REGION Network 4: Run IGG Sea Water P301-CV311-CV322
   // Changed to 560 from 580
   RUNG wire#powerrail
      { S7_Templates := "SrcType := Int" } GE_Contact(in1 := "100_GCU_AUTO_SEQ_DB".CRNT_STEP, in2 := 50)
      { S7_Templates := "SrcType := Int" } LE_Contact(in1 := "100_GCU_AUTO_SEQ_DB".CRNT_STEP, in2 := 560)
      wire#w1
      Contact( "51_SLAVE_STATUS".CV322_OPN )
      Contact( "51_SLAVE_STATUS"."CV-321_CLSD" )
      Coil( "56_SLAVE_CMNDS".OPEN_CV311 )
   END_RUNG
   RUNG wire#powerrail
      I_Contact( "10_DI_DATA".E_400_STPD )
      I_Contact( "10_DI_DATA".E_400_SHTDN )
   END_RUNG wire#w1
   RUNG wire#w1
      Coil( "56_SLAVE_CMNDS".OPEN_CV322 )
   END_RUNG
   RUNG wire#w1
      Contact( "51_SLAVE_STATUS".CV311_OPN )
      Contact( "51_SLAVE_STATUS".CV322_OPN )
      Coil( "56_SLAVE_CMNDS".RUN_P301 )
   END_RUNG
   // the same network as SCL:
   #_w1 := (("100_GCU_AUTO_SEQ_DB".CRNT_STEP >= 50) AND ("100_GCU_AUTO_SEQ_DB".CRNT_STEP <= 560)) OR (NOT "10_DI_DATA".E_400_STPD AND NOT "10_DI_DATA".E_400_SHTDN);
   "56_SLAVE_CMNDS".OPEN_CV311 := #_w1 AND "51_SLAVE_STATUS".CV322_OPN AND "51_SLAVE_STATUS"."CV-321_CLSD";
   "56_SLAVE_CMNDS".OPEN_CV322 := #_w1;
   "56_SLAVE_CMNDS".RUN_P301 := #_w1 AND "51_SLAVE_STATUS".CV311_OPN AND "51_SLAVE_STATUS".CV322_OPN;
END_REGION

REGION Network 5: Q136.0 - Fresh Water Fill Valve Control(CV358)
   // True = RUN, False = NOT
   RUNG wire#powerrail
      { S7_Templates := "SrcType := Int" } GE_Contact(in1 := "100_GCU_AUTO_SEQ_DB".CRNT_STEP, in2 := 90)
      { S7_Templates := "SrcType := Int" } LT_Contact(in1 := "100_GCU_AUTO_SEQ_DB".CRNT_STEP, in2 := 200)
      wire#w1
      Coil( "14_DQ_DATA".CV_358 )
   END_RUNG
   RUNG wire#powerrail
      Contact( "108_GCU_TNK_REFILL_SEQ_DB".OPEN_CV358 )
   END_RUNG wire#w1
   RUNG wire#powerrail
      Contact( "110_GCU_TNK_FLUSH_SEQ_DB".OPEN_CV358 )
   END_RUNG wire#w1
   // the same network as SCL:
   "14_DQ_DATA".CV_358 := (("100_GCU_AUTO_SEQ_DB".CRNT_STEP >= 90) AND ("100_GCU_AUTO_SEQ_DB".CRNT_STEP < 200)) OR "108_GCU_TNK_REFILL_SEQ_DB".OPEN_CV358 OR "110_GCU_TNK_FLUSH_SEQ_DB".OPEN_CV358;
END_REGION

REGION Network 6: Q136.1 - Waste Water Drain Valve Control (CV341)
   // True = Close, False = Open    Condition added to avoid back filling the GCU through common drain on Bordeira
   RUNG wire#powerrail
      { S7_Templates := "SrcType := Int" } GE_Contact(in1 := "100_GCU_AUTO_SEQ_DB".CRNT_STEP, in2 := 60)
      { S7_Templates := "SrcType := Int" } LT_Contact(in1 := "100_GCU_AUTO_SEQ_DB".CRNT_STEP, in2 := 570)
      wire#w1
      Coil( "14_DQ_DATA".CV_341 )
   END_RUNG
   RUNG wire#powerrail
      I_Contact( "51_SLAVE_STATUS".CV311_CLSD )
      Contact( "AlwaysTRUE" )
   END_RUNG wire#w1
   // the same network as SCL:
   "14_DQ_DATA".CV_341 := (("100_GCU_AUTO_SEQ_DB".CRNT_STEP >= 60) AND ("100_GCU_AUTO_SEQ_DB".CRNT_STEP < 570)) OR (NOT "51_SLAVE_STATUS".CV311_CLSD AND "AlwaysTRUE");
END_REGION

REGION Network 7: Q136.2 - Block Valve 1 Control (CV407) +++Control By BWTS+++
   // True = RUN, False = NOT
END_REGION

REGION Network 8: Q136.3 - Bleed Valve Control (CV409) +++Control By BWTS+++
   // True = OPEN, False = CLOSE
END_REGION

REGION Network 9: Q136.4 - Block Valve 2 Control (CV411) +++Control By BWTS+++
   // True = OPEN, False = CLOSE
END_REGION

REGION Network 10: Q136.5 - Ambient Air Valve Control (CV441)
   // True = CLOSE, False = OPEN        STOP bits are redundant.
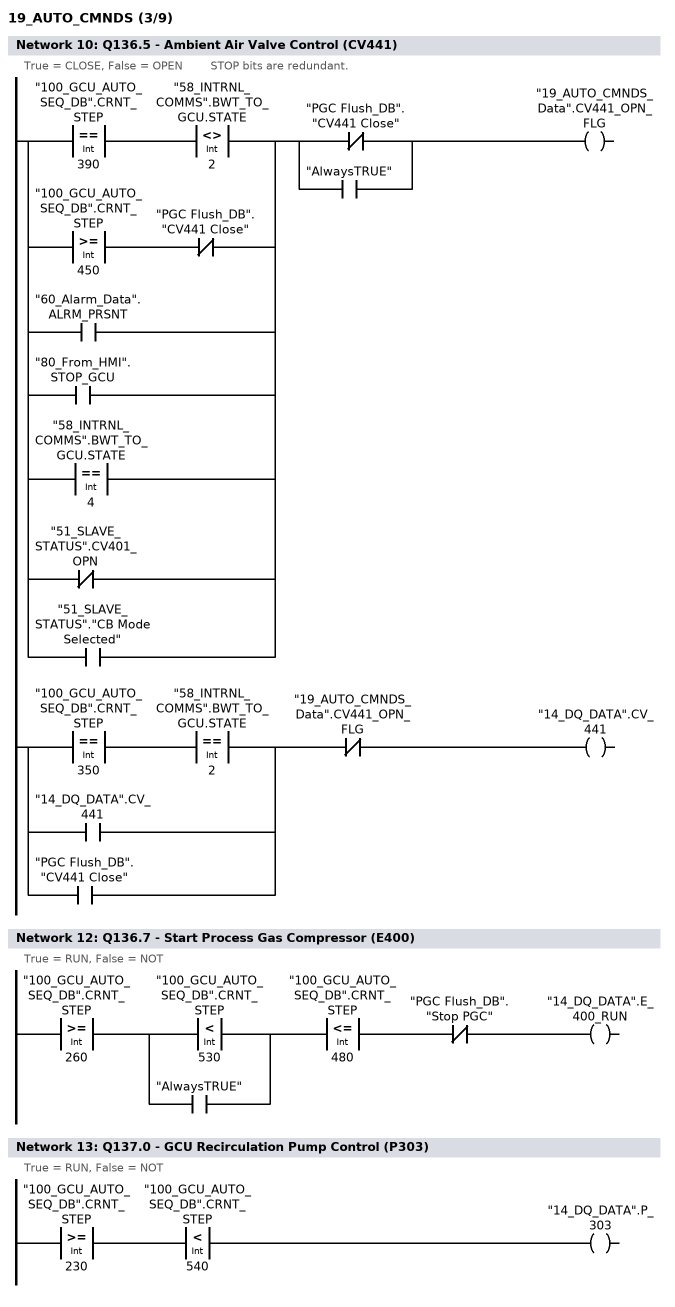
   RUNG wire#powerrail
      { S7_Templates := "SrcType := Int" } EQ_Contact(in1 := "100_GCU_AUTO_SEQ_DB".CRNT_STEP, in2 := 390)
      { S7_Templates := "SrcType := Int" } NE_Contact(in1 := "58_INTRNL_COMMS".BWT_TO_GCU.STATE, in2 := 2)
      wire#w1
      I_Contact( "PGC Flush_DB"."CV441 Close" )
      wire#w2
      Coil( "19_AUTO_CMNDS_Data".CV441_OPN_FLG )
   END_RUNG
   RUNG wire#powerrail
      { S7_Templates := "SrcType := Int" } GE_Contact(in1 := "100_GCU_AUTO_SEQ_DB".CRNT_STEP, in2 := 450)
      I_Contact( "PGC Flush_DB"."CV441 Close" )
   END_RUNG wire#w1
   RUNG wire#powerrail
      Contact( "60_Alarm_Data".ALRM_PRSNT )
   END_RUNG wire#w1
   RUNG wire#powerrail
      Contact( "80_From_HMI".STOP_GCU )
   END_RUNG wire#w1
   RUNG wire#powerrail
      { S7_Templates := "SrcType := Int" } EQ_Contact(in1 := "58_INTRNL_COMMS".BWT_TO_GCU.STATE, in2 := 4)
   END_RUNG wire#w1
   RUNG wire#powerrail
      I_Contact( "51_SLAVE_STATUS".CV401_OPN )
   END_RUNG wire#w1
   RUNG wire#powerrail
      Contact( "51_SLAVE_STATUS"."CB Mode Selected" )
   END_RUNG wire#w1
   RUNG wire#w1
      Contact( "AlwaysTRUE" )
   END_RUNG wire#w2
   RUNG wire#powerrail
      { S7_Templates := "SrcType := Int" } EQ_Contact(in1 := "100_GCU_AUTO_SEQ_DB".CRNT_STEP, in2 := 350)
      { S7_Templates := "SrcType := Int" } EQ_Contact(in1 := "58_INTRNL_COMMS".BWT_TO_GCU.STATE, in2 := 2)
      wire#w3
      I_Contact( "19_AUTO_CMNDS_Data".CV441_OPN_FLG )
      Coil( "14_DQ_DATA".CV_441 )
   END_RUNG
   RUNG wire#powerrail
      Contact( "14_DQ_DATA".CV_441 )
   END_RUNG wire#w3
   RUNG wire#powerrail
      Contact( "PGC Flush_DB"."CV441 Close" )
   END_RUNG wire#w3
   // the same network as SCL:
   "19_AUTO_CMNDS_Data".CV441_OPN_FLG := ((("100_GCU_AUTO_SEQ_DB".CRNT_STEP = 390) AND ("58_INTRNL_COMMS".BWT_TO_GCU.STATE <> 2)) OR (("100_GCU_AUTO_SEQ_DB".CRNT_STEP >= 450) AND NOT "PGC Flush_DB"."CV441 Close") OR "60_Alarm_Data".ALRM_PRSNT OR "80_From_HMI".STOP_GCU OR ("58_INTRNL_COMMS".BWT_TO_GCU.STATE = 4) OR NOT "51_SLAVE_STATUS".CV401_OPN OR "51_SLAVE_STATUS"."CB Mode Selected") AND (NOT "PGC Flush_DB"."CV441 Close" OR "AlwaysTRUE");
   "14_DQ_DATA".CV_441 := ((("100_GCU_AUTO_SEQ_DB".CRNT_STEP = 350) AND ("58_INTRNL_COMMS".BWT_TO_GCU.STATE = 2)) OR "14_DQ_DATA".CV_441 OR "PGC Flush_DB"."CV441 Close") AND NOT "19_AUTO_CMNDS_Data".CV441_OPN_FLG;
END_REGION

REGION Network 11: Q136.6 - Main Gas to Deck Valve Control (CV406) +++Control By BWTS+++
   // True = RUN, False = NOT
END_REGION

REGION Network 12: Q136.7 - Start Process Gas Compressor (E400)
   // True = RUN, False = NOT
   RUNG wire#powerrail
      { S7_Templates := "SrcType := Int" } GE_Contact(in1 := "100_GCU_AUTO_SEQ_DB".CRNT_STEP, in2 := 260)
      wire#w1
      { S7_Templates := "SrcType := Int" } LT_Contact(in1 := "100_GCU_AUTO_SEQ_DB".CRNT_STEP, in2 := 530)
      wire#w2
      { S7_Templates := "SrcType := Int" } LE_Contact(in1 := "100_GCU_AUTO_SEQ_DB".CRNT_STEP, in2 := 480)
      I_Contact( "PGC Flush_DB"."Stop PGC" )
      Coil( "14_DQ_DATA".E_400_RUN )
   END_RUNG
   RUNG wire#w1
      Contact( "AlwaysTRUE" )
   END_RUNG wire#w2
   // the same network as SCL:
   "14_DQ_DATA".E_400_RUN := ("100_GCU_AUTO_SEQ_DB".CRNT_STEP >= 260) AND (("100_GCU_AUTO_SEQ_DB".CRNT_STEP < 530) OR "AlwaysTRUE") AND ("100_GCU_AUTO_SEQ_DB".CRNT_STEP <= 480) AND NOT "PGC Flush_DB"."Stop PGC";
END_REGION

REGION Network 13: Q137.0 - GCU Recirculation Pump Control (P303)
   // True = RUN, False = NOT
   RUNG wire#powerrail
      { S7_Templates := "SrcType := Int" } GE_Contact(in1 := "100_GCU_AUTO_SEQ_DB".CRNT_STEP, in2 := 230)
      { S7_Templates := "SrcType := Int" } LT_Contact(in1 := "100_GCU_AUTO_SEQ_DB".CRNT_STEP, in2 := 540)
      Coil( "14_DQ_DATA".P_303 )
   END_RUNG
   // the same network as SCL:
   "14_DQ_DATA".P_303 := ("100_GCU_AUTO_SEQ_DB".CRNT_STEP >= 230) AND ("100_GCU_AUTO_SEQ_DB".CRNT_STEP < 540);
END_REGION

REGION Network 14: Q137.1 - GCU Booster Pump Control (P304)
   // True = ALARM, False = NOT
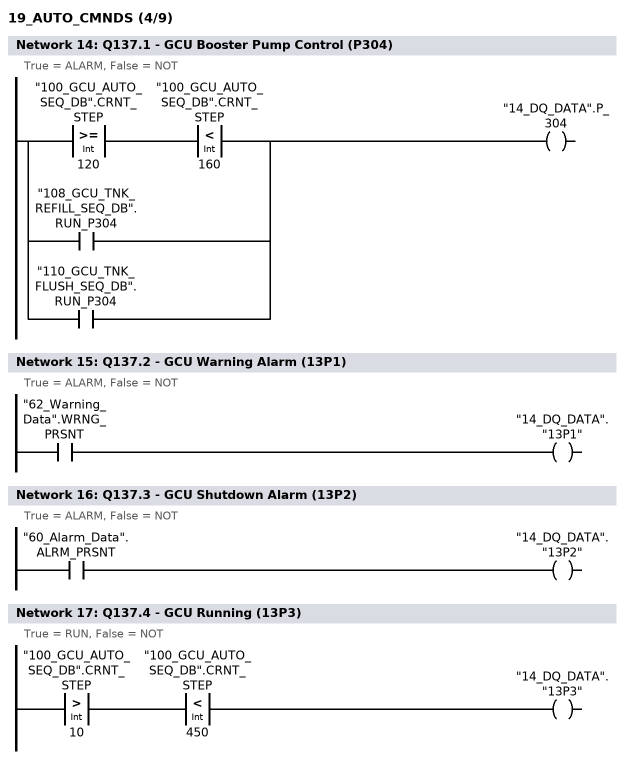
   RUNG wire#powerrail
      { S7_Templates := "SrcType := Int" } GE_Contact(in1 := "100_GCU_AUTO_SEQ_DB".CRNT_STEP, in2 := 120)
      { S7_Templates := "SrcType := Int" } LT_Contact(in1 := "100_GCU_AUTO_SEQ_DB".CRNT_STEP, in2 := 160)
      wire#w1
      Coil( "14_DQ_DATA".P_304 )
   END_RUNG
   RUNG wire#powerrail
      Contact( "108_GCU_TNK_REFILL_SEQ_DB".RUN_P304 )
   END_RUNG wire#w1
   RUNG wire#powerrail
      Contact( "110_GCU_TNK_FLUSH_SEQ_DB".RUN_P304 )
   END_RUNG wire#w1
   // the same network as SCL:
   "14_DQ_DATA".P_304 := (("100_GCU_AUTO_SEQ_DB".CRNT_STEP >= 120) AND ("100_GCU_AUTO_SEQ_DB".CRNT_STEP < 160)) OR "108_GCU_TNK_REFILL_SEQ_DB".RUN_P304 OR "110_GCU_TNK_FLUSH_SEQ_DB".RUN_P304;
END_REGION

REGION Network 15: Q137.2 - GCU Warning Alarm (13P1)
   // True = ALARM, False = NOT
   RUNG wire#powerrail
      Contact( "62_Warning_Data".WRNG_PRSNT )
      Coil( "14_DQ_DATA"."13P1" )
   END_RUNG
   // the same network as SCL:
   "14_DQ_DATA"."13P1" := "62_Warning_Data".WRNG_PRSNT;
END_REGION

REGION Network 16: Q137.3 - GCU Shutdown Alarm (13P2)
   // True = ALARM, False = NOT
   RUNG wire#powerrail
      Contact( "60_Alarm_Data".ALRM_PRSNT )
      Coil( "14_DQ_DATA"."13P2" )
   END_RUNG
   // the same network as SCL:
   "14_DQ_DATA"."13P2" := "60_Alarm_Data".ALRM_PRSNT;
END_REGION

REGION Network 17: Q137.4 - GCU Running (13P3)
   // True = RUN, False = NOT
   RUNG wire#powerrail
      { S7_Templates := "SrcType := Int" } GT_Contact(in1 := "100_GCU_AUTO_SEQ_DB".CRNT_STEP, in2 := 10)
      { S7_Templates := "SrcType := Int" } LT_Contact(in1 := "100_GCU_AUTO_SEQ_DB".CRNT_STEP, in2 := 450)
      Coil( "14_DQ_DATA"."13P3" )
   END_RUNG
   // the same network as SCL:
   "14_DQ_DATA"."13P3" := ("100_GCU_AUTO_SEQ_DB".CRNT_STEP > 10) AND ("100_GCU_AUTO_SEQ_DB".CRNT_STEP < 450);
END_REGION

REGION Network 18: Q137.5 - Ballast Water Tank Level HI HI (13P4)
   // True = ALARM, False = NOT
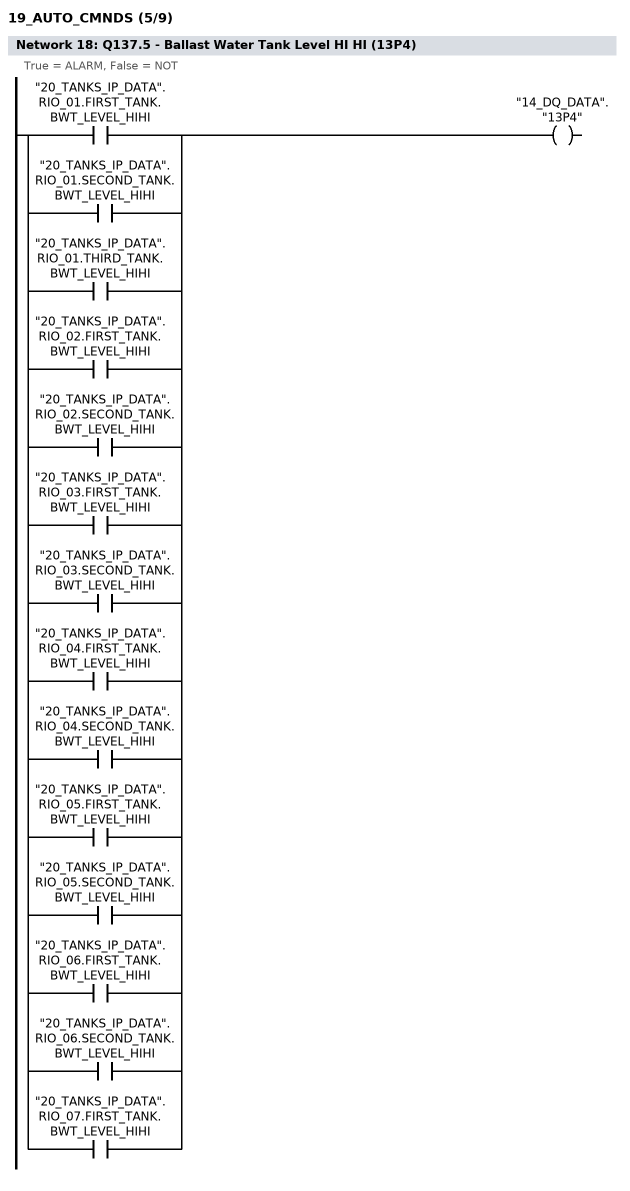
   RUNG wire#powerrail
      Contact( "20_TANKS_IP_DATA".RIO_01.FIRST_TANK.BWT_LEVEL_HIHI )
      wire#w1
      Coil( "14_DQ_DATA"."13P4" )
   END_RUNG
   RUNG wire#powerrail
      Contact( "20_TANKS_IP_DATA".RIO_01.SECOND_TANK.BWT_LEVEL_HIHI )
   END_RUNG wire#w1
   RUNG wire#powerrail
      Contact( "20_TANKS_IP_DATA".RIO_01.THIRD_TANK.BWT_LEVEL_HIHI )
   END_RUNG wire#w1
   RUNG wire#powerrail
      Contact( "20_TANKS_IP_DATA".RIO_02.FIRST_TANK.BWT_LEVEL_HIHI )
   END_RUNG wire#w1
   RUNG wire#powerrail
      Contact( "20_TANKS_IP_DATA".RIO_02.SECOND_TANK.BWT_LEVEL_HIHI )
   END_RUNG wire#w1
   RUNG wire#powerrail
      Contact( "20_TANKS_IP_DATA".RIO_03.FIRST_TANK.BWT_LEVEL_HIHI )
   END_RUNG wire#w1
   RUNG wire#powerrail
      Contact( "20_TANKS_IP_DATA".RIO_03.SECOND_TANK.BWT_LEVEL_HIHI )
   END_RUNG wire#w1
   RUNG wire#powerrail
      Contact( "20_TANKS_IP_DATA".RIO_04.FIRST_TANK.BWT_LEVEL_HIHI )
   END_RUNG wire#w1
   RUNG wire#powerrail
      Contact( "20_TANKS_IP_DATA".RIO_04.SECOND_TANK.BWT_LEVEL_HIHI )
   END_RUNG wire#w1
   RUNG wire#powerrail
      Contact( "20_TANKS_IP_DATA".RIO_05.FIRST_TANK.BWT_LEVEL_HIHI )
   END_RUNG wire#w1
   RUNG wire#powerrail
      Contact( "20_TANKS_IP_DATA".RIO_05.SECOND_TANK.BWT_LEVEL_HIHI )
   END_RUNG wire#w1
   RUNG wire#powerrail
      Contact( "20_TANKS_IP_DATA".RIO_06.FIRST_TANK.BWT_LEVEL_HIHI )
   END_RUNG wire#w1
   RUNG wire#powerrail
      Contact( "20_TANKS_IP_DATA".RIO_06.SECOND_TANK.BWT_LEVEL_HIHI )
   END_RUNG wire#w1
   RUNG wire#powerrail
      Contact( "20_TANKS_IP_DATA".RIO_07.FIRST_TANK.BWT_LEVEL_HIHI )
   END_RUNG wire#w1
   // the same network as SCL:
   "14_DQ_DATA"."13P4" := "20_TANKS_IP_DATA".RIO_01.FIRST_TANK.BWT_LEVEL_HIHI OR "20_TANKS_IP_DATA".RIO_01.SECOND_TANK.BWT_LEVEL_HIHI OR "20_TANKS_IP_DATA".RIO_01.THIRD_TANK.BWT_LEVEL_HIHI OR "20_TANKS_IP_DATA".RIO_02.FIRST_TANK.BWT_LEVEL_HIHI OR "20_TANKS_IP_DATA".RIO_02.SECOND_TANK.BWT_LEVEL_HIHI OR "20_TANKS_IP_DATA".RIO_03.FIRST_TANK.BWT_LEVEL_HIHI OR "20_TANKS_IP_DATA".RIO_03.SECOND_TANK.BWT_LEVEL_HIHI OR "20_TANKS_IP_DATA".RIO_04.FIRST_TANK.BWT_LEVEL_HIHI OR "20_TANKS_IP_DATA".RIO_04.SECOND_TANK.BWT_LEVEL_HIHI OR "20_TANKS_IP_DATA".RIO_05.FIRST_TANK.BWT_LEVEL_HIHI OR "20_TANKS_IP_DATA".RIO_05.SECOND_TANK.BWT_LEVEL_HIHI OR "20_TANKS_IP_DATA".RIO_06.FIRST_TANK.BWT_LEVEL_HIHI OR "20_TANKS_IP_DATA".RIO_06.SECOND_TANK.BWT_LEVEL_HIHI OR "20_TANKS_IP_DATA".RIO_07.FIRST_TANK.BWT_LEVEL_HIHI;
END_REGION

REGION Network 19: Q137.6 - GCU Alarm Buzzer (13P5)
   // True = ALARM, False = NOT
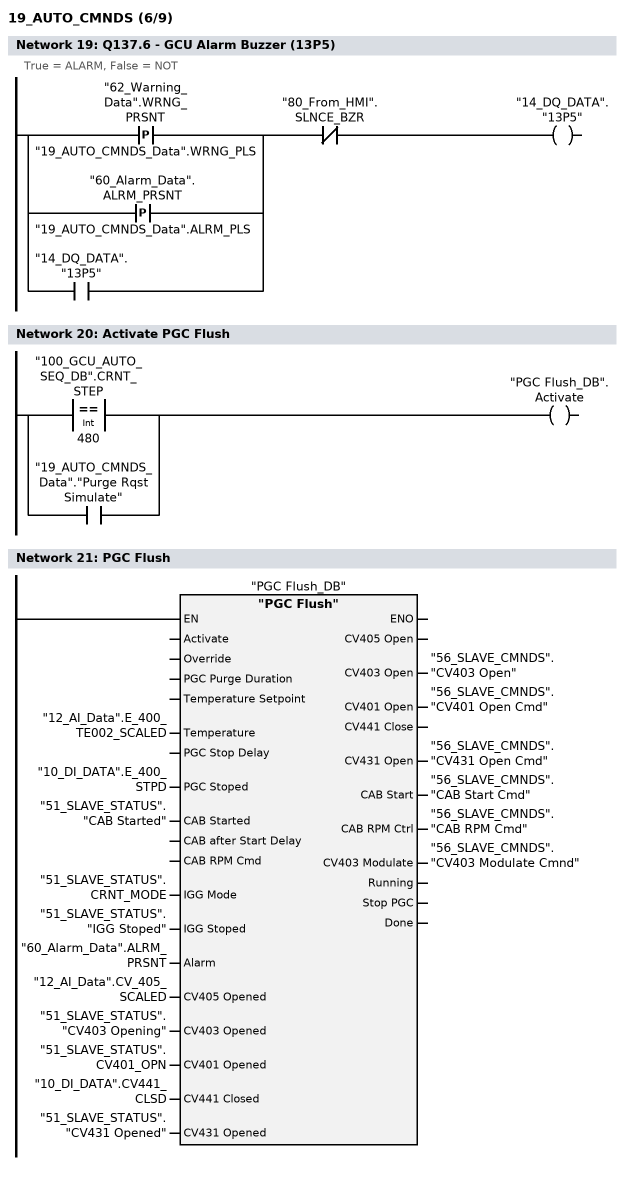
   RUNG wire#powerrail
      P_Contact(operand := "62_Warning_Data".WRNG_PRSNT, bit := "19_AUTO_CMNDS_Data".WRNG_PLS)
      wire#w1
      I_Contact( "80_From_HMI".SLNCE_BZR )
      Coil( "14_DQ_DATA"."13P5" )
   END_RUNG
   RUNG wire#powerrail
      P_Contact(operand := "60_Alarm_Data".ALRM_PRSNT, bit := "19_AUTO_CMNDS_Data".ALRM_PLS)
   END_RUNG wire#w1
   RUNG wire#powerrail
      Contact( "14_DQ_DATA"."13P5" )
   END_RUNG wire#w1
   // the same network as SCL:
   #_w1 := "62_Warning_Data".WRNG_PRSNT AND NOT "19_AUTO_CMNDS_Data".WRNG_PLS;   // rising edge of "62_Warning_Data".WRNG_PRSNT
   "19_AUTO_CMNDS_Data".WRNG_PLS := "62_Warning_Data".WRNG_PRSNT;
   #_w2 := "60_Alarm_Data".ALRM_PRSNT AND NOT "19_AUTO_CMNDS_Data".ALRM_PLS;   // rising edge of "60_Alarm_Data".ALRM_PRSNT
   "19_AUTO_CMNDS_Data".ALRM_PLS := "60_Alarm_Data".ALRM_PRSNT;
   "14_DQ_DATA"."13P5" := (#_w1 OR #_w2 OR "14_DQ_DATA"."13P5") AND NOT "80_From_HMI".SLNCE_BZR;
END_REGION

REGION Network 20: Activate PGC Flush
   RUNG wire#powerrail
      { S7_Templates := "SrcType := Int" } EQ_Contact(in1 := "100_GCU_AUTO_SEQ_DB".CRNT_STEP, in2 := 480)
      wire#w1
      Coil( "PGC Flush_DB".Activate )
   END_RUNG
   RUNG wire#powerrail
      Contact( "19_AUTO_CMNDS_Data"."Purge Rqst Simulate" )
   END_RUNG wire#w1
   // the same network as SCL:
   "PGC Flush_DB".Activate := ("100_GCU_AUTO_SEQ_DB".CRNT_STEP = 480) OR "19_AUTO_CMNDS_Data"."Purge Rqst Simulate";
END_REGION

REGION Network 21: PGC Flush
   RUNG wire#powerrail
      "PGC Flush_DB"(Activate :=, Override :=, "PGC Purge Duration" :=, "Temperature Setpoint" :=, Temperature := "12_AI_Data".E_400_TE002_SCALED, "PGC Stop Delay" :=, "PGC Stoped" := "10_DI_DATA".E_400_STPD, "CAB Started" := "51_SLAVE_STATUS"."CAB Started", "CAB after Start Delay" :=, "CAB RPM Cmd" :=, "IGG Mode" := "51_SLAVE_STATUS".CRNT_MODE, "IGG Stoped" := "51_SLAVE_STATUS"."IGG Stoped", Alarm := "60_Alarm_Data".ALRM_PRSNT, "CV405 Opened" := "12_AI_Data".CV_405_SCALED, "CV403 Opened" := "51_SLAVE_STATUS"."CV403 Opening", "CV401 Opened" := "51_SLAVE_STATUS".CV401_OPN, "CV441 Closed" := "10_DI_DATA".CV441_CLSD, "CV431 Opened" := "51_SLAVE_STATUS"."CV431 Opened", "CV405 Open" =>, "CV403 Open" => "56_SLAVE_CMNDS"."CV403 Open", "CV401 Open" => "56_SLAVE_CMNDS"."CV401 Open Cmd", "CV441 Close" =>, "CV431 Open" => "56_SLAVE_CMNDS"."CV431 Open Cmd", "CAB Start" => "56_SLAVE_CMNDS"."CAB Start Cmd", "CAB RPM Ctrl" => "56_SLAVE_CMNDS"."CAB RPM Cmd", "CV403 Modulate" => "56_SLAVE_CMNDS"."CV403 Modulate Cmnd", Running =>, "Stop PGC" =>, Done =>)
   END_RUNG
   // the same network as SCL:
   "PGC Flush_DB"(Temperature := "12_AI_Data".E_400_TE002_SCALED,   // "PGC Flush"
                  "PGC Stoped" := "10_DI_DATA".E_400_STPD,
                  "CAB Started" := "51_SLAVE_STATUS"."CAB Started",
                  "IGG Mode" := "51_SLAVE_STATUS".CRNT_MODE,
                  "IGG Stoped" := "51_SLAVE_STATUS"."IGG Stoped",
                  Alarm := "60_Alarm_Data".ALRM_PRSNT,
                  "CV405 Opened" := "12_AI_Data".CV_405_SCALED,
                  "CV403 Opened" := "51_SLAVE_STATUS"."CV403 Opening",
                  "CV401 Opened" := "51_SLAVE_STATUS".CV401_OPN,
                  "CV441 Closed" := "10_DI_DATA".CV441_CLSD,
                  "CV431 Opened" := "51_SLAVE_STATUS"."CV431 Opened",
                  "CV403 Open" => "56_SLAVE_CMNDS"."CV403 Open",
                  "CV401 Open" => "56_SLAVE_CMNDS"."CV401 Open Cmd",
                  "CV431 Open" => "56_SLAVE_CMNDS"."CV431 Open Cmd",
                  "CAB Start" => "56_SLAVE_CMNDS"."CAB Start Cmd",
                  "CAB RPM Ctrl" => "56_SLAVE_CMNDS"."CAB RPM Cmd",
                  "CV403 Modulate" => "56_SLAVE_CMNDS"."CV403 Modulate Cmnd");
END_REGION

REGION Network 22: Q137.7 - Stop Process Gas Compressor (E400)
   // True = ALARM, False = NOT
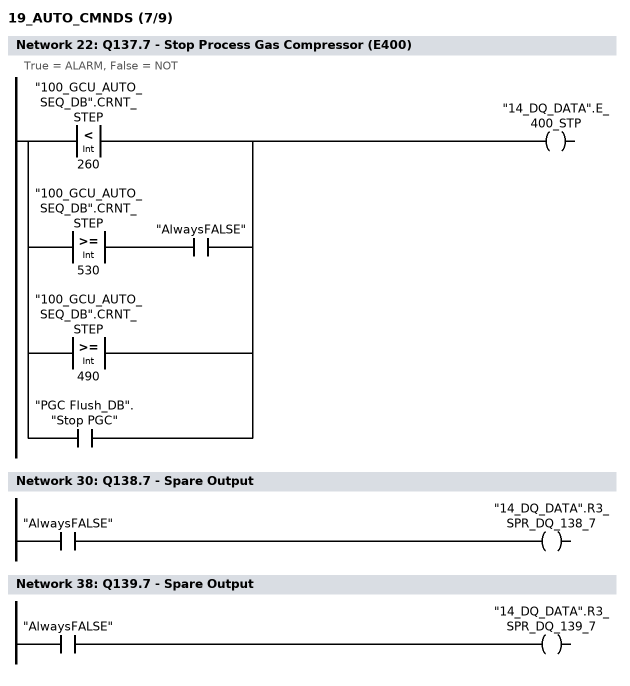
   RUNG wire#powerrail
      { S7_Templates := "SrcType := Int" } LT_Contact(in1 := "100_GCU_AUTO_SEQ_DB".CRNT_STEP, in2 := 260)
      wire#w1
      Coil( "14_DQ_DATA".E_400_STP )
   END_RUNG
   RUNG wire#powerrail
      { S7_Templates := "SrcType := Int" } GE_Contact(in1 := "100_GCU_AUTO_SEQ_DB".CRNT_STEP, in2 := 530)
      Contact( "AlwaysFALSE" )
   END_RUNG wire#w1
   RUNG wire#powerrail
      { S7_Templates := "SrcType := Int" } GE_Contact(in1 := "100_GCU_AUTO_SEQ_DB".CRNT_STEP, in2 := 490)
   END_RUNG wire#w1
   RUNG wire#powerrail
      Contact( "PGC Flush_DB"."Stop PGC" )
   END_RUNG wire#w1
   // the same network as SCL:
   "14_DQ_DATA".E_400_STP := ("100_GCU_AUTO_SEQ_DB".CRNT_STEP < 260) OR (("100_GCU_AUTO_SEQ_DB".CRNT_STEP >= 530) AND "AlwaysFALSE") OR ("100_GCU_AUTO_SEQ_DB".CRNT_STEP >= 490) OR "PGC Flush_DB"."Stop PGC";
END_REGION

REGION Network 23: Q138.0 - Pilot For GTT FPT Valve (CV422-FPT) +++Control By BWTS+++
END_REGION

REGION Network 24: Q138.1 - Pilot For GTT 1 Port Valve (CV422-1P) +++Control By BWTS+++
END_REGION

REGION Network 25: Q138.2 - Pilot For GTT 1 Starboard Valve (CV421-1S) +++Control By BWTS+++
END_REGION

REGION Network 26: Q138.3 - Pilot For GTT 2 Port Valve (CV422-2P) +++Control By BWTS+++
END_REGION

REGION Network 27: Q138.4 - Pilot For GTT 2 Starboard Valve (CV421-2S) +++Control By BWTS+++
END_REGION

REGION Network 28: Q138.5 - Pilot For GTT 3 Port Valve (CV422-3P) +++Control By BWTS+++
END_REGION

REGION Network 29: Q138.6 - Pilot For GTT 3 Starboard Valve (CV421-3S) +++Control By BWTS+++
END_REGION

REGION Network 30: Q138.7 - Spare Output
   RUNG wire#powerrail
      Contact( "AlwaysFALSE" )
      Coil( "14_DQ_DATA".R3_SPR_DQ_138_7 )
   END_RUNG
   // the same network as SCL:
   "14_DQ_DATA".R3_SPR_DQ_138_7 := "AlwaysFALSE";
END_REGION

REGION Network 31: Q139.0 - Pilot For GTT 4 Port Valve (CV422-4P) +++Control By BWTS+++
END_REGION

REGION Network 32: Q139.1 - Pilot For GTT 4 Starboard Valve (CV421-4S) +++Control By BWTS+++
END_REGION

REGION Network 33: Q139.2 - Pilot For GTT 5 Port Valve (CV422-5P) +++Control By BWTS+++
END_REGION

REGION Network 34: Q139.3 - Pilot For GTT 5 Starboard Valve (CV421-5S) +++Control By BWTS+++
END_REGION

REGION Network 35: Q139.4 - Pilot For GTT 6 Port Valve (CV422-6P) +++Control By BWTS+++
END_REGION

REGION Network 36: Q139.5 - Pilot For GTT 6 Starboard Valve (CV421-6S) +++Control By BWTS+++
END_REGION

REGION Network 37: Q139.6 - Pilot For GTT APT Valve (CV422-APT) +++Control By BWTS+++
END_REGION

REGION Network 38: Q139.7 - Spare Output
   RUNG wire#powerrail
      Contact( "AlwaysFALSE" )
      Coil( "14_DQ_DATA".R3_SPR_DQ_139_7 )
   END_RUNG
   // the same network as SCL:
   "14_DQ_DATA".R3_SPR_DQ_139_7 := "AlwaysFALSE";
END_REGION

REGION Network 39: QW800 - CV405 Gas Vent Position Control
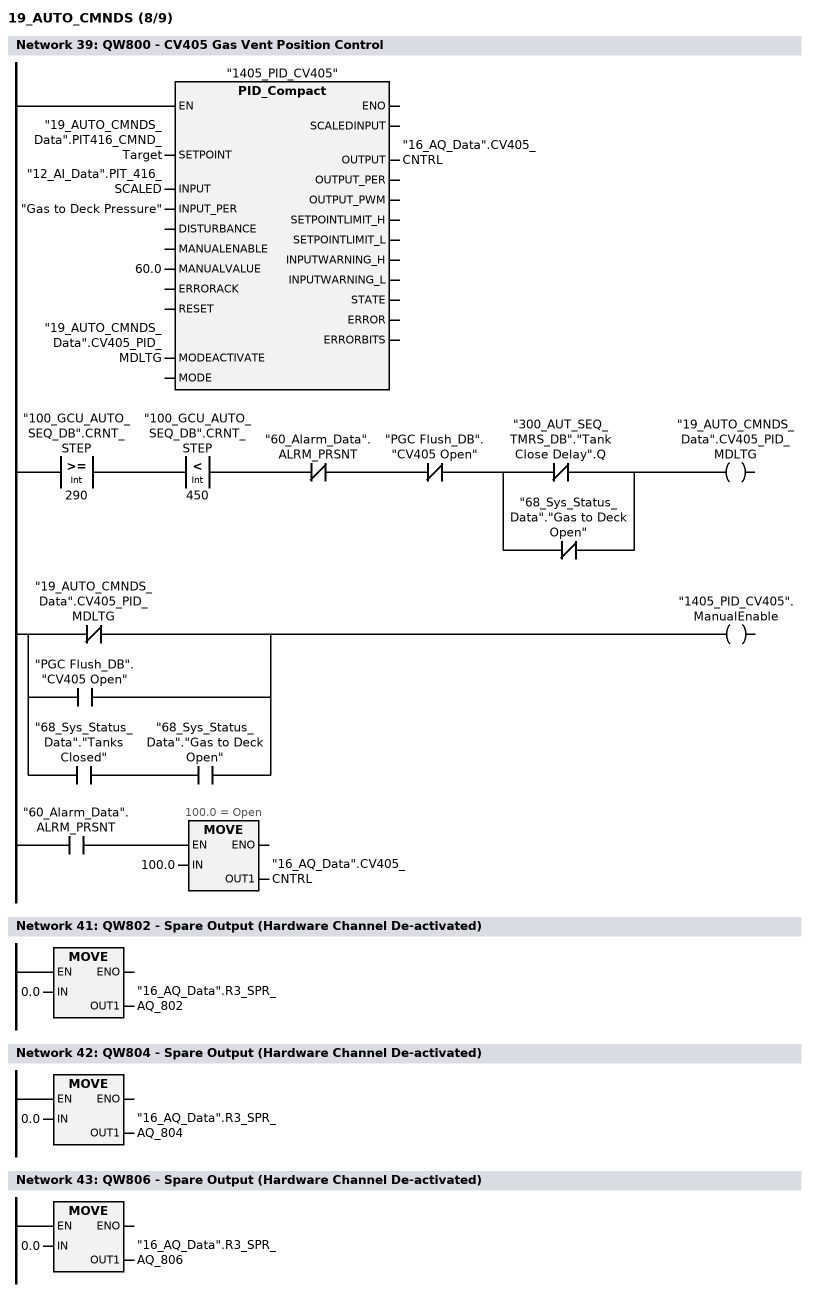
   "1405_PID_CV405"(Setpoint := "19_AUTO_CMNDS_Data".PIT416_CMND_Target,   // PID_Compact
                    Input := "12_AI_Data".PIT_416_SCALED,
                    Input_PER := "Gas to Deck Pressure",
                    ManualValue := 60.0,
                    ModeActivate := "19_AUTO_CMNDS_Data".CV405_PID_MDLTG,
                    Output => "16_AQ_Data".CV405_CNTRL);
   "19_AUTO_CMNDS_Data".CV405_PID_MDLTG := ("100_GCU_AUTO_SEQ_DB".CRNT_STEP >= 290) AND ("100_GCU_AUTO_SEQ_DB".CRNT_STEP < 450) AND NOT "60_Alarm_Data".ALRM_PRSNT AND NOT "PGC Flush_DB"."CV405 Open" AND (NOT "300_AUT_SEQ_TMRS_DB"."Tank Close Delay".Q OR NOT "68_Sys_Status_Data"."Gas to Deck Open");
   "1405_PID_CV405".ManualEnable := NOT "19_AUTO_CMNDS_Data".CV405_PID_MDLTG OR "PGC Flush_DB"."CV405 Open" OR ("68_Sys_Status_Data"."Tanks Closed" AND "68_Sys_Status_Data"."Gas to Deck Open");
   IF "60_Alarm_Data".ALRM_PRSNT THEN
       "16_AQ_Data".CV405_CNTRL := 100.0;   // 100.0 = Open
   END_IF;
END_REGION

REGION Network 41: QW802 - Spare Output (Hardware Channel De-activated)
   RUNG wire#powerrail
      Move(in := 0.0, out1 => "16_AQ_Data".R3_SPR_AQ_802)
   END_RUNG
   // the same network as SCL:
   "16_AQ_Data".R3_SPR_AQ_802 := 0.0;
END_REGION

REGION Network 42: QW804 - Spare Output (Hardware Channel De-activated)
   RUNG wire#powerrail
      Move(in := 0.0, out1 => "16_AQ_Data".R3_SPR_AQ_804)
   END_RUNG
   // the same network as SCL:
   "16_AQ_Data".R3_SPR_AQ_804 := 0.0;
END_REGION

REGION Network 43: QW806 - Spare Output (Hardware Channel De-activated)
   RUNG wire#powerrail
      Move(in := 0.0, out1 => "16_AQ_Data".R3_SPR_AQ_806)
   END_RUNG
   // the same network as SCL:
   "16_AQ_Data".R3_SPR_AQ_806 := 0.0;
END_REGION

REGION Network 44: Run Command To IGG
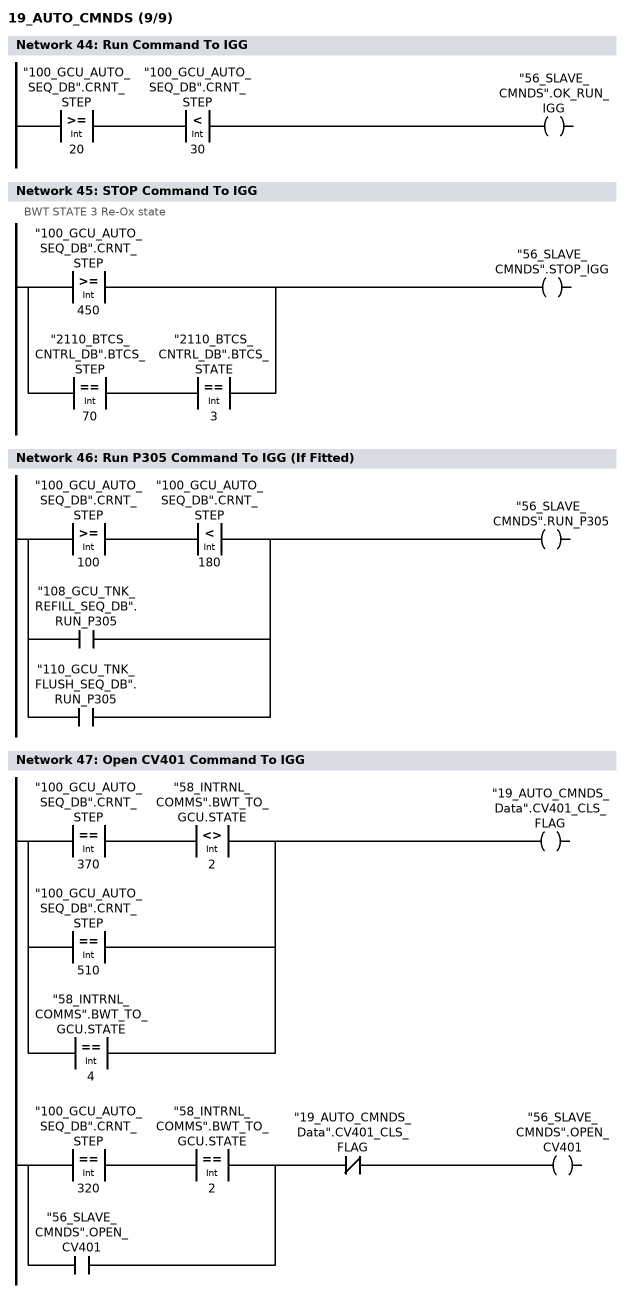
   RUNG wire#powerrail
      { S7_Templates := "SrcType := Int" } GE_Contact(in1 := "100_GCU_AUTO_SEQ_DB".CRNT_STEP, in2 := 20)
      { S7_Templates := "SrcType := Int" } LT_Contact(in1 := "100_GCU_AUTO_SEQ_DB".CRNT_STEP, in2 := 30)
      Coil( "56_SLAVE_CMNDS".OK_RUN_IGG )
   END_RUNG
   // the same network as SCL:
   "56_SLAVE_CMNDS".OK_RUN_IGG := ("100_GCU_AUTO_SEQ_DB".CRNT_STEP >= 20) AND ("100_GCU_AUTO_SEQ_DB".CRNT_STEP < 30);
END_REGION

REGION Network 45: STOP Command To IGG
   // BWT STATE 3 Re-Ox state
   RUNG wire#powerrail
      { S7_Templates := "SrcType := Int" } GE_Contact(in1 := "100_GCU_AUTO_SEQ_DB".CRNT_STEP, in2 := 450)
      wire#w1
      Coil( "56_SLAVE_CMNDS".STOP_IGG )
   END_RUNG
   RUNG wire#powerrail
      { S7_Templates := "SrcType := Int" } EQ_Contact(in1 := "2110_BTCS_CNTRL_DB".BTCS_STEP, in2 := 70)
      { S7_Templates := "SrcType := Int" } EQ_Contact(in1 := "2110_BTCS_CNTRL_DB".BTCS_STATE, in2 := 3)
   END_RUNG wire#w1
   // the same network as SCL:
   "56_SLAVE_CMNDS".STOP_IGG := ("100_GCU_AUTO_SEQ_DB".CRNT_STEP >= 450) OR (("2110_BTCS_CNTRL_DB".BTCS_STEP = 70) AND ("2110_BTCS_CNTRL_DB".BTCS_STATE = 3));
END_REGION

REGION Network 46: Run P305 Command To IGG (If Fitted)
   RUNG wire#powerrail
      { S7_Templates := "SrcType := Int" } GE_Contact(in1 := "100_GCU_AUTO_SEQ_DB".CRNT_STEP, in2 := 100)
      { S7_Templates := "SrcType := Int" } LT_Contact(in1 := "100_GCU_AUTO_SEQ_DB".CRNT_STEP, in2 := 180)
      wire#w1
      Coil( "56_SLAVE_CMNDS".RUN_P305 )
   END_RUNG
   RUNG wire#powerrail
      Contact( "108_GCU_TNK_REFILL_SEQ_DB".RUN_P305 )
   END_RUNG wire#w1
   RUNG wire#powerrail
      Contact( "110_GCU_TNK_FLUSH_SEQ_DB".RUN_P305 )
   END_RUNG wire#w1
   // the same network as SCL:
   "56_SLAVE_CMNDS".RUN_P305 := (("100_GCU_AUTO_SEQ_DB".CRNT_STEP >= 100) AND ("100_GCU_AUTO_SEQ_DB".CRNT_STEP < 180)) OR "108_GCU_TNK_REFILL_SEQ_DB".RUN_P305 OR "110_GCU_TNK_FLUSH_SEQ_DB".RUN_P305;
END_REGION

REGION Network 47: Open CV401 Command To IGG
   RUNG wire#powerrail
      { S7_Templates := "SrcType := Int" } EQ_Contact(in1 := "100_GCU_AUTO_SEQ_DB".CRNT_STEP, in2 := 370)
      { S7_Templates := "SrcType := Int" } NE_Contact(in1 := "58_INTRNL_COMMS".BWT_TO_GCU.STATE, in2 := 2)
      wire#w1
      Coil( "19_AUTO_CMNDS_Data".CV401_CLS_FLAG )
   END_RUNG
   RUNG wire#powerrail
      { S7_Templates := "SrcType := Int" } EQ_Contact(in1 := "100_GCU_AUTO_SEQ_DB".CRNT_STEP, in2 := 510)
   END_RUNG wire#w1
   RUNG wire#powerrail
      { S7_Templates := "SrcType := Int" } EQ_Contact(in1 := "58_INTRNL_COMMS".BWT_TO_GCU.STATE, in2 := 4)
   END_RUNG wire#w1
   RUNG wire#powerrail
      { S7_Templates := "SrcType := Int" } EQ_Contact(in1 := "100_GCU_AUTO_SEQ_DB".CRNT_STEP, in2 := 320)
      { S7_Templates := "SrcType := Int" } EQ_Contact(in1 := "58_INTRNL_COMMS".BWT_TO_GCU.STATE, in2 := 2)
      wire#w2
      I_Contact( "19_AUTO_CMNDS_Data".CV401_CLS_FLAG )
      Coil( "56_SLAVE_CMNDS".OPEN_CV401 )
   END_RUNG
   RUNG wire#powerrail
      Contact( "56_SLAVE_CMNDS".OPEN_CV401 )
   END_RUNG wire#w2
   // the same network as SCL:
   "19_AUTO_CMNDS_Data".CV401_CLS_FLAG := (("100_GCU_AUTO_SEQ_DB".CRNT_STEP = 370) AND ("58_INTRNL_COMMS".BWT_TO_GCU.STATE <> 2)) OR ("100_GCU_AUTO_SEQ_DB".CRNT_STEP = 510) OR ("58_INTRNL_COMMS".BWT_TO_GCU.STATE = 4);
   "56_SLAVE_CMNDS".OPEN_CV401 := ((("100_GCU_AUTO_SEQ_DB".CRNT_STEP = 320) AND ("58_INTRNL_COMMS".BWT_TO_GCU.STATE = 2)) OR "56_SLAVE_CMNDS".OPEN_CV401) AND NOT "19_AUTO_CMNDS_Data".CV401_CLS_FLAG;
END_REGION
END_FUNCTION

// folder: 100 - 199 Automatic Sequencing

FUNCTION_BLOCK "100_GCU_AUTO_SEQ"   // FB100, LAD
TITLE = Automatic Sequence
{ S7_Optimized_Access := 'TRUE' }
AUTHOR : JRS
VERSION : 0.1
// Master sequencing for automatic operation
   VAR_INPUT
      RST : Bool;   // Sequence reset
   END_VAR
   VAR_OUTPUT
      RNG : Bool;   // Sequence running
   END_VAR
   VAR
      CRNT_STEP : Int;
      STEP_001 : "500_SEQ_STEP";
      STEP_005 : "500_SEQ_STEP";
      STEP_010 : "500_SEQ_STEP";
      STEP_020 : "500_SEQ_STEP";
      STEP_030 : "500_SEQ_STEP";
      STEP_040 : "500_SEQ_STEP";
      STEP_050 : "500_SEQ_STEP";
      STEP_060 : "500_SEQ_STEP";
      STEP_070 : "500_SEQ_STEP";
      STEP_080 : "500_SEQ_STEP";
      STEP_090 : "500_SEQ_STEP";
      STEP_100 : "500_SEQ_STEP";
      STEP_110 : "500_SEQ_STEP";
      STEP_120 : "500_SEQ_STEP";
      STEP_130 : "500_SEQ_STEP";
      STEP_140 : "500_SEQ_STEP";
      STEP_150 : "500_SEQ_STEP";
      STEP_160 : "500_SEQ_STEP";
      STEP_170 : "500_SEQ_STEP";
      STEP_180 : "500_SEQ_STEP";
      STEP_190 : "500_SEQ_STEP";
      STEP_200 : "500_SEQ_STEP";
      STEP_210 : "500_SEQ_STEP";
      STEP_220 : "500_SEQ_STEP";
      STEP_230 : "500_SEQ_STEP";
      STEP_240 : "500_SEQ_STEP";
      STEP_250 : "500_SEQ_STEP";
      STEP_260 : "500_SEQ_STEP";
      STEP_270 : "500_SEQ_STEP";
      STEP_280 : "500_SEQ_STEP";
      STEP_290 : "500_SEQ_STEP";
      STEP_300 : "500_SEQ_STEP";
      STEP_310 : "500_SEQ_STEP";
      STEP_320 : "500_SEQ_STEP";
      STEP_330 : "500_SEQ_STEP";
      STEP_340 : "500_SEQ_STEP";
      STEP_350 : "500_SEQ_STEP";
      STEP_360 : "500_SEQ_STEP";
      STEP_370 : "500_SEQ_STEP";
      STEP_380 : "500_SEQ_STEP";
      STEP_390 : "500_SEQ_STEP";
      STEP_400 : "500_SEQ_STEP";
      STEP_410 : "500_SEQ_STEP";
      STEP_420 : "500_SEQ_STEP";
      STEP_430 : "500_SEQ_STEP";
      STEP_440 : "500_SEQ_STEP";
      STEP_450 : "500_SEQ_STEP";
      STEP_460 : "500_SEQ_STEP";
      STEP_470 : "500_SEQ_STEP";
      STEP_480 : "500_SEQ_STEP";
      STEP_490 : "500_SEQ_STEP";
      STEP_500 : "500_SEQ_STEP";
      STEP_510 : "500_SEQ_STEP";
      STEP_520 : "500_SEQ_STEP";
      STEP_530 : "500_SEQ_STEP";
      STEP_540 : "500_SEQ_STEP";
      STEP_550 : "500_SEQ_STEP";
      STEP_560 : "500_SEQ_STEP";
      STEP_570 : "500_SEQ_STEP";
      STEP_580 : "500_SEQ_STEP";
      STEP_590 : "500_SEQ_STEP";
      STEP_600 : "500_SEQ_STEP";
      STEP_610 : "500_SEQ_STEP";
      STEP_620 : "500_SEQ_STEP";
      STEP_630 : "500_SEQ_STEP";
   END_VAR
   VAR_TEMP   // added for the SCL form of the ladder/FBD networks
      _w1 : Bool;
      _w2 : Bool;
   END_VAR
BEGIN

REGION Network 1: Auto Initiated or Reset = Set Step to 0
   // Going into automatic or sequence reset resets the sequence
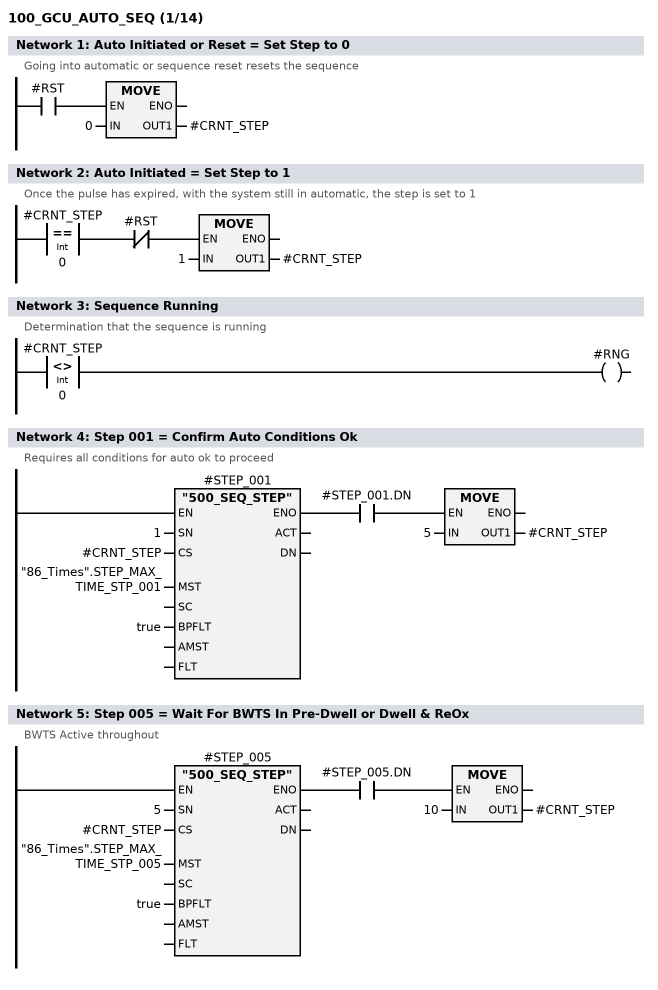
   RUNG wire#powerrail
      Contact( #RST )
      Move(in := 0, out1 => #CRNT_STEP)
   END_RUNG
   // the same network as SCL:
   IF #RST THEN #CRNT_STEP := 0; END_IF;
END_REGION
